       "R-201_Write_TO_T-101_DB".Abort := "R-201_SEQ_DB".S_NO >= 21 AND "R-201_SEQ_DB".S_NO <= 39;
       "R-201_Write_TO_T-102_DB".Abort := "R-201_SEQ_DB".S_NO >= 21 AND "R-201_SEQ_DB".S_NO <= 39;
       "R-201_Write_TO_T-103_DB".Abort :=("R-201_DB".Status.State = 3);

   END_IF;

   //***************Interlocks to T-104***************//
   "R-201_Write_TO_T-104_DB".ReqWater := "XV-2013_DB".CS AND "XV-1043_DB".OS AND ("R-201_DB".Status.Step = 23 OR "R-201_DB".Status.Step = 68 OR "R-201_DB".Status.Step = 66);

   //***************Valves Status***************//
   "R-201_Aux_DB"."Bool".TOff := "R-201_DB".Equipments.Valves."XV-2013".TurningOff OR "R-201_DB".Equipments.Valves."XV-2011".TurningOff OR "R-201_DB".Equipments.Valves."XV-2021".TurningOff OR "R-201_DB".Equipments.Valves."XV-1043".TurningOff;

   //***************Timers***************//
   //Pre-Mix Timer
   "R-201_Aux_DB"."Bool".PreMixT_En := "R-201_DB".Status.Step = 26 AND "R-201_Read_FROM_T-102_DB".Recirculating AND "R-201_Read_FROM_T-101_DB".Recirculating; //T-102 AND T-102 Mixing
   "R-201_Aux_DB"."Bool".PreMixT_Reset := "R-201_DB".Cmds.Abort OR "R-201_DB".Status.Step = 1;
   //pH Stabilize Timer
   "R-201_Aux_DB"."Bool".StabpHTEn := "R-201_Aux_DB"."Bool".StabpHTEnStep AND "FT-1021_DB".SAI > 0.1 AND "FT-1011_DB".SAI > 0.1;
   "R-201_Aux_DB"."Bool".StabpHTEn_Reset := "R-201_DB".Cmds.Abort OR "R-201_DB".Status.Step = 1;
   //Reaction Timer
   "R-201_Aux_DB"."Bool".ReactorTEn := "R-201_DB".Status.Step = 40;
   "R-201_Aux_DB"."Bool".ReactorT_Reset := "R-201_DB".Cmds.Abort OR "R-201_DB".Status.Step = 1;
   //Last Run Timer
   "R-201_Aux_DB"."Bool".FlushOutTEn := ("R-201_DB".Status.Step = 67 OR "R-201_DB".Status.Step = 64) AND ("P-201A_DB".CF OR "P-201B_DB".CF) AND "XV-2013_DB".OS;
   //Mix To Clean Timer
   "R-201_Aux_DB"."Bool".MixToCleanTEn := "R-201_DB".Status.Step = 63 AND "VFD-R201_DB".RUN_FEEDBACK;
   "R-201_Aux_DB"."Bool".MixToCleanT_Reset := "R-201_DB".Cmds.Abort OR "R-201_DB".Status.Step = 1;
END_FUNCTION

FUNCTION "R-201_SEQ_FC" : Void   // FC37, LAD
{ S7_Optimized_Access := 'TRUE' }
VERSION : 0.1
   VAR_TEMP   // added for the SCL form of the ladder/FBD networks
      _w1 : Bool;
      _w2 : Bool;
   END_VAR
BEGIN

REGION Network 2: Abort
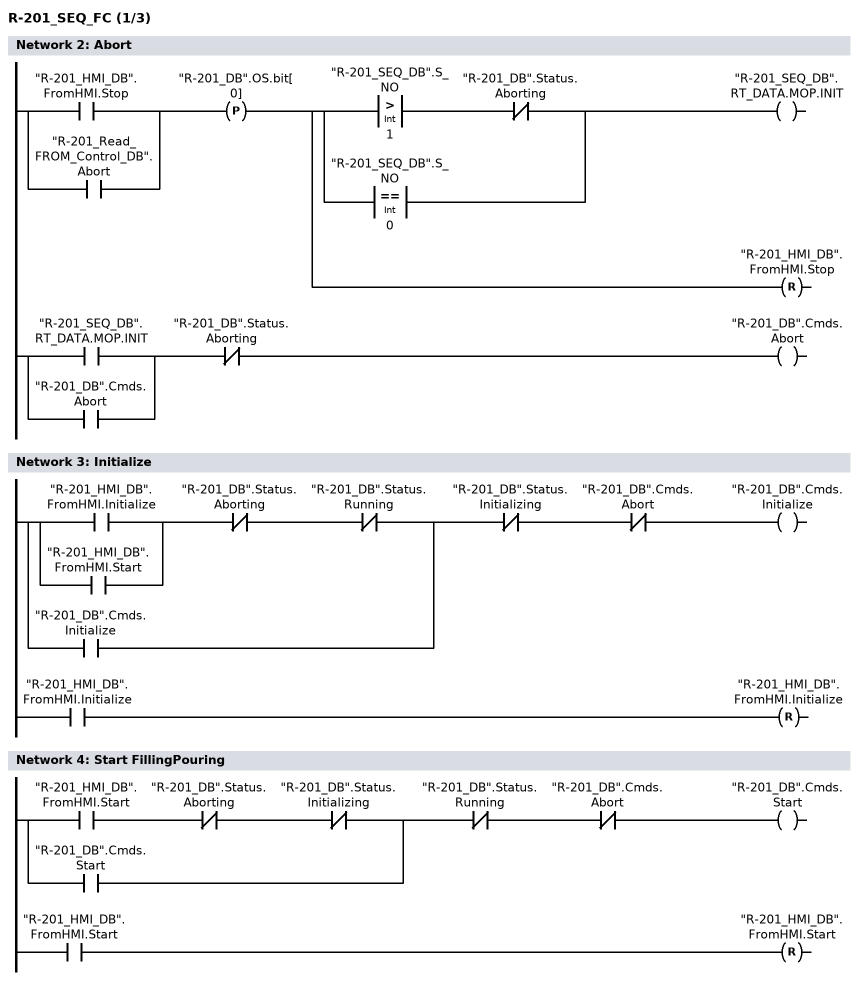
   RUNG wire#powerrail
      Contact( "R-201_HMI_DB".FromHMI.Stop )
      wire#w1
      P_Trig( "R-201_DB".OS.bit[0] )
      wire#w2
      { S7_Templates := "SrcType := Int" } GT_Contact(in1 := "R-201_SEQ_DB".S_NO, in2 := 1)
      I_Contact( "R-201_DB".Status.Aborting )
      wire#w3
      Coil( "R-201_SEQ_DB".RT_DATA.MOP.INIT )
   END_RUNG
   RUNG wire#powerrail
      Contact( "R-201_Read_FROM_Control_DB".Abort )
   END_RUNG wire#w1
   RUNG wire#w2
      { S7_Templates := "SrcType := Int" } EQ_Contact(in1 := "R-201_SEQ_DB".S_NO, in2 := 0)
   END_RUNG wire#w3
   RUNG wire#w2
      R_Coil( "R-201_HMI_DB".FromHMI.Stop )
   END_RUNG
   RUNG wire#powerrail
      Contact( "R-201_SEQ_DB".RT_DATA.MOP.INIT )
      wire#w4
      I_Contact( "R-201_DB".Status.Aborting )
      Coil( "R-201_DB".Cmds.Abort )
   END_RUNG
   RUNG wire#powerrail
      Contact( "R-201_DB".Cmds.Abort )
   END_RUNG wire#w4
   // the same network as SCL:
   #_w1 := "R-201_HMI_DB".FromHMI.Stop OR "R-201_Read_FROM_Control_DB".Abort;
   #_w2 := #_w1 AND NOT "R-201_DB".OS.bit[0];   // rising edge
   "R-201_DB".OS.bit[0] := #_w1;
   "R-201_SEQ_DB".RT_DATA.MOP.INIT := #_w2 AND ((("R-201_SEQ_DB".S_NO > 1) AND NOT "R-201_DB".Status.Aborting) OR ("R-201_SEQ_DB".S_NO = 0));
   IF #_w2 THEN "R-201_HMI_DB".FromHMI.Stop := FALSE; END_IF;
   "R-201_DB".Cmds.Abort := ("R-201_SEQ_DB".RT_DATA.MOP.INIT OR "R-201_DB".Cmds.Abort) AND NOT "R-201_DB".Status.Aborting;
END_REGION

REGION Network 3: Initialize
   RUNG wire#powerrail
      Contact( "R-201_HMI_DB".FromHMI.Initialize )
      wire#w1
      I_Contact( "R-201_DB".Status.Aborting )
      I_Contact( "R-201_DB".Status.Running )
      wire#w2
      I_Contact( "R-201_DB".Status.Initializing )
      I_Contact( "R-201_DB".Cmds.Abort )
      Coil( "R-201_DB".Cmds.Initialize )
   END_RUNG
   RUNG wire#powerrail
      Contact( "R-201_HMI_DB".FromHMI.Start )
   END_RUNG wire#w1
   RUNG wire#powerrail
      Contact( "R-201_DB".Cmds.Initialize )
   END_RUNG wire#w2
   RUNG wire#powerrail
      Contact( "R-201_HMI_DB".FromHMI.Initialize )
      R_Coil( "R-201_HMI_DB".FromHMI.Initialize )
   END_RUNG
   // the same network as SCL:
   "R-201_DB".Cmds.Initialize := ((("R-201_HMI_DB".FromHMI.Initialize OR "R-201_HMI_DB".FromHMI.Start) AND NOT "R-201_DB".Status.Aborting AND NOT "R-201_DB".Status.Running) OR "R-201_DB".Cmds.Initialize) AND NOT "R-201_DB".Status.Initializing AND NOT "R-201_DB".Cmds.Abort;
   IF "R-201_HMI_DB".FromHMI.Initialize THEN "R-201_HMI_DB".FromHMI.Initialize := FALSE; END_IF;
END_REGION

REGION Network 4: Start FillingPouring
   RUNG wire#powerrail
      Contact( "R-201_HMI_DB".FromHMI.Start )
      I_Contact( "R-201_DB".Status.Aborting )
      I_Contact( "R-201_DB".Status.Initializing )
      wire#w1
      I_Contact( "R-201_DB".Status.Running )
      I_Contact( "R-201_DB".Cmds.Abort )
      Coil( "R-201_DB".Cmds.Start )
   END_RUNG
   RUNG wire#powerrail
      Contact( "R-201_DB".Cmds.Start )
   END_RUNG wire#w1
   RUNG wire#powerrail
      Contact( "R-201_HMI_DB".FromHMI.Start )
      R_Coil( "R-201_HMI_DB".FromHMI.Start )
   END_RUNG
   // the same network as SCL:
   "R-201_DB".Cmds.Start := (("R-201_HMI_DB".FromHMI.Start AND NOT "R-201_DB".Status.Aborting AND NOT "R-201_DB".Status.Initializing) OR "R-201_DB".Cmds.Start) AND NOT "R-201_DB".Status.Running AND NOT "R-201_DB".Cmds.Abort;
   IF "R-201_HMI_DB".FromHMI.Start THEN "R-201_HMI_DB".FromHMI.Start := FALSE; END_IF;
END_REGION

REGION Network 5: Procedure Selected
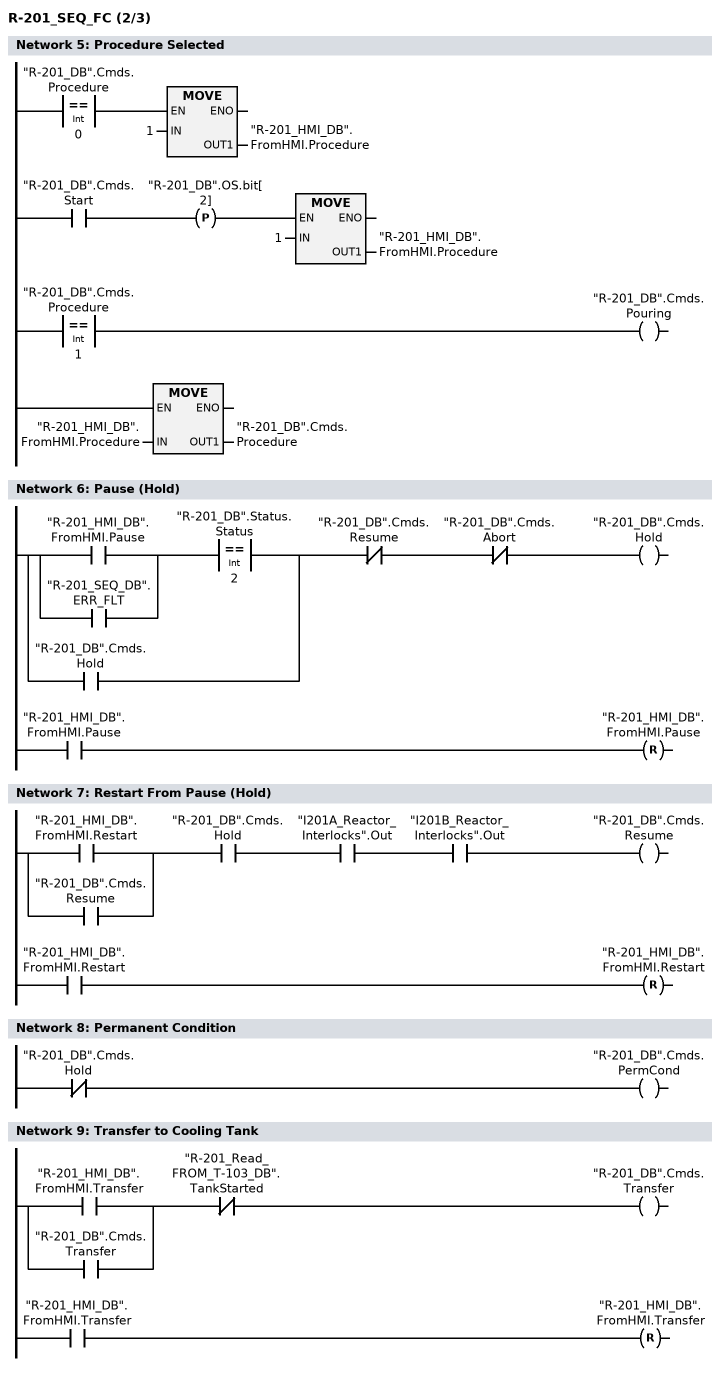
   RUNG wire#powerrail
      { S7_Templates := "SrcType := Int" } EQ_Contact(in1 := "R-201_DB".Cmds.Procedure, in2 := 0)
      Move(in := 1, out1 => "R-201_HMI_DB".FromHMI.Procedure)
   END_RUNG
   RUNG wire#powerrail
      Contact( "R-201_DB".Cmds.Start )
      P_Trig( "R-201_DB".OS.bit[2] )
      Move(in := 1, out1 => "R-201_HMI_DB".FromHMI.Procedure)
   END_RUNG
   RUNG wire#powerrail
      { S7_Templates := "SrcType := Int" } EQ_Contact(in1 := "R-201_DB".Cmds.Procedure, in2 := 1)
      Coil( "R-201_DB".Cmds.Pouring )
   END_RUNG
   RUNG wire#powerrail
      Move(in := "R-201_HMI_DB".FromHMI.Procedure, out1 => "R-201_DB".Cmds.Procedure)
   END_RUNG
   // the same network as SCL:
   IF "R-201_DB".Cmds.Procedure = 0 THEN "R-201_HMI_DB".FromHMI.Procedure := 1; END_IF;
   #_w1 := "R-201_DB".Cmds.Start AND NOT "R-201_DB".OS.bit[2];   // rising edge
   "R-201_DB".OS.bit[2] := "R-201_DB".Cmds.Start;
   IF #_w1 THEN "R-201_HMI_DB".FromHMI.Procedure := 1; END_IF;
   "R-201_DB".Cmds.Pouring := "R-201_DB".Cmds.Procedure = 1;
   "R-201_DB".Cmds.Procedure := "R-201_HMI_DB".FromHMI.Procedure;
END_REGION

REGION Network 6: Pause (Hold)
   RUNG wire#powerrail
      Contact( "R-201_HMI_DB".FromHMI.Pause )
      wire#w1
      { S7_Templates := "SrcType := Int" } EQ_Contact(in1 := "R-201_DB".Status.Status, in2 := 2)
      wire#w2
      I_Contact( "R-201_DB".Cmds.Resume )
      I_Contact( "R-201_DB".Cmds.Abort )
      Coil( "R-201_DB".Cmds.Hold )
   END_RUNG
   RUNG wire#powerrail
      Contact( "R-201_SEQ_DB".ERR_FLT )
   END_RUNG wire#w1
   RUNG wire#powerrail
      Contact( "R-201_DB".Cmds.Hold )
   END_RUNG wire#w2
   RUNG wire#powerrail
      Contact( "R-201_HMI_DB".FromHMI.Pause )
      R_Coil( "R-201_HMI_DB".FromHMI.Pause )
   END_RUNG
   // the same network as SCL:
   "R-201_DB".Cmds.Hold := ((("R-201_HMI_DB".FromHMI.Pause OR "R-201_SEQ_DB".ERR_FLT) AND ("R-201_DB".Status.Status = 2)) OR "R-201_DB".Cmds.Hold) AND NOT "R-201_DB".Cmds.Resume AND NOT "R-201_DB".Cmds.Abort;
   IF "R-201_HMI_DB".FromHMI.Pause THEN "R-201_HMI_DB".FromHMI.Pause := FALSE; END_IF;
END_REGION

REGION Network 7: Restart From Pause (Hold)
   RUNG wire#powerrail
      Contact( "R-201_HMI_DB".FromHMI.Restart )
      wire#w1
      Contact( "R-201_DB".Cmds.Hold )
      Contact( "I201A_Reactor_Interlocks".Out )
      Contact( "I201B_Reactor_Interlocks".Out )
      Coil( "R-201_DB".Cmds.Resume )
   END_RUNG
   RUNG wire#powerrail
      Contact( "R-201_DB".Cmds.Resume )
   END_RUNG wire#w1
   RUNG wire#powerrail
      Contact( "R-201_HMI_DB".FromHMI.Restart )
      R_Coil( "R-201_HMI_DB".FromHMI.Restart )
   END_RUNG
   // the same network as SCL:
   "R-201_DB".Cmds.Resume := ("R-201_HMI_DB".FromHMI.Restart OR "R-201_DB".Cmds.Resume) AND "R-201_DB".Cmds.Hold AND "I201A_Reactor_Interlocks".Out AND "I201B_Reactor_Interlocks".Out;
   IF "R-201_HMI_DB".FromHMI.Restart THEN "R-201_HMI_DB".FromHMI.Restart := FALSE; END_IF;
END_REGION

REGION Network 8: Permanent Condition
   RUNG wire#powerrail
      I_Contact( "R-201_DB".Cmds.Hold )
      Coil( "R-201_DB".Cmds.PermCond )
   END_RUNG
   // the same network as SCL:
   "R-201_DB".Cmds.PermCond := NOT "R-201_DB".Cmds.Hold;
END_REGION

REGION Network 9: Transfer to Cooling Tank
   RUNG wire#powerrail
      Contact( "R-201_HMI_DB".FromHMI.Transfer )
      wire#w1
      I_Contact( "R-201_Read_FROM_T-103_DB".TankStarted )
      Coil( "R-201_DB".Cmds.Transfer )
   END_RUNG
   RUNG wire#powerrail
      Contact( "R-201_DB".Cmds.Transfer )
   END_RUNG wire#w1
   RUNG wire#powerrail
      Contact( "R-201_HMI_DB".FromHMI.Transfer )
      R_Coil( "R-201_HMI_DB".FromHMI.Transfer )
   END_RUNG
   // the same network as SCL:
   "R-201_DB".Cmds.Transfer := ("R-201_HMI_DB".FromHMI.Transfer OR "R-201_DB".Cmds.Transfer) AND NOT "R-201_Read_FROM_T-103_DB".TankStarted;
   IF "R-201_HMI_DB".FromHMI.Transfer THEN "R-201_HMI_DB".FromHMI.Transfer := FALSE; END_IF;
END_REGION

REGION Network 10: Tank Wash
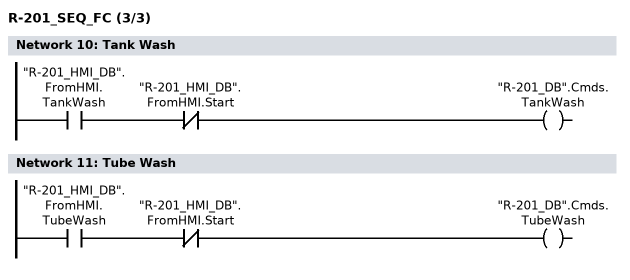
   RUNG wire#powerrail
      Contact( "R-201_HMI_DB".FromHMI.TankWash )
      I_Contact( "R-201_HMI_DB".FromHMI.Start )
      Coil( "R-201_DB".Cmds.TankWash )
   END_RUNG
   // the same network as SCL:
   "R-201_DB".Cmds.TankWash := "R-201_HMI_DB".FromHMI.TankWash AND NOT "R-201_HMI_DB".FromHMI.Start;
END_REGION

REGION Network 11: Tube Wash
   RUNG wire#powerrail
      Contact( "R-201_HMI_DB".FromHMI.TubeWash )
      I_Contact( "R-201_HMI_DB".FromHMI.Start )
      Coil( "R-201_DB".Cmds.TubeWash )
   END_RUNG
   // the same network as SCL:
   "R-201_DB".Cmds.TubeWash := "R-201_HMI_DB".FromHMI.TubeWash AND NOT "R-201_HMI_DB".FromHMI.Start;
END_REGION

REGION Network 12 (SCL): Sequence Status
   IF "R-201_SEQ_DB".S_NO = 1 THEN
       "R-201_DB".Status.Status := 1; //Idle
   ELSIF ("R-201_SEQ_DB".S_NO > 1 AND "R-201_SEQ_DB".S_NO <= 150)  AND NOT "R-201_SEQ_DB".ERR_FLT AND NOT "R-201_DB".Cmds.Hold THEN
       "R-201_DB".Status.Status := 2; //Running
   ELSIF "R-201_SEQ_DB".S_NO >= 151 AND "R-201_SEQ_DB".S_NO <= 160 AND NOT "R-201_SEQ_DB".ERR_FLT THEN
       "R-201_DB".Status.Status := 3; // Stopping
   ELSIF "R-201_SEQ_DB".ERR_FLT  AND ("R-201_SEQ_DB".S_NO > 1 AND "R-201_SEQ_DB".S_NO <= 150) THEN
       "R-201_DB".Status.Status := 4; //Held
   ELSIF "R-201_SEQ_DB".ERR_FLT AND  ("R-201_SEQ_DB".S_NO > 1 AND "R-201_SEQ_DB".S_NO <= 150) AND "R-201_Aux_DB"."Bool".TOff  THEN
       "R-201_DB".Status.Status := 5; // Holding
   ELSE
       "R-201_DB".Status.Status := 6; // Unknown
   END_IF;


   "R-201_DB".Status.Running := ("R-201_SEQ_DB".S_NO > 3 AND "R-201_SEQ_DB".S_NO <= 150);
   "R-201_DB".Status.Initializing := ("R-201_SEQ_DB".S_NO >= 141 AND "R-201_SEQ_DB".S_NO <= 150);
   //Enable/Disable HMI Start/Stop Button
   "R-201_HMI_DB".ToHMI.EnStopButton:=("R-201_DB".Status.Status>1) OR "R-201_DB".Status.Step=0; //Enable HMI Stop Button
   "R-201_HMI_DB".ToHMI.EnStartButton:= "R-201_DB".Status.Status = 1; //Enable Start Button
   "R-201_HMI_DB".ToHMI.EnPauseButton := "R-201_DB".Status.Status = 2; //Enable Pause Button
   "R-201_HMI_DB".ToHMI.EnRestartButton := "R-201_DB".Status.Status = 4; //Enable Restart Button

   //****Interlock Activated
   "R-201_HMI_DB".ToHMI.InterlockActivated := "I201A_Reactor_Interlocks".Out AND "I201B_Reactor_Interlocks".Out;
END_REGION

REGION Network 13 (SCL): Sequence Step
   "R-201_DB".Status.Step := "R-201_SEQ_DB".S_NO;
END_REGION

REGION Network 14 (SCL): Sequence state (Procedure running)
   IF "R-201_SEQ_DB".S_NO = 3 OR "R-201_SEQ_DB".S_NO = 4 THEN
       "R-201_DB".Status.State := 1; //Seq Selection
   ELSIF "R-201_SEQ_DB".S_NO >= 21 AND "R-201_SEQ_DB".S_NO <= 60 THEN
       "R-201_DB".Status.State := 2; //Pouring 
   ELSIF "R-201_SEQ_DB".S_NO >= 61 AND "R-201_SEQ_DB".S_NO <= 80 THEN
       "R-201_DB".Status.State := 3; //Transfering
   ELSIF "R-201_SEQ_DB".S_NO >= 81 AND "R-201_SEQ_DB".S_NO <= 100 THEN
       "R-201_DB".Status.State := 4; //Washing Tank
   ELSIF "R-201_SEQ_DB".S_NO >= 101 AND "R-201_SEQ_DB".S_NO <= 140 THEN
       "R-201_DB".Status.State := 5; //Washing Lines
   ELSIF "R-201_SEQ_DB".S_NO >= 151 AND "R-201_SEQ_DB".S_NO <= 160 THEN
       "R-201_DB".Status.State := 6; //Aborting
   ELSIF "R-201_SEQ_DB".S_NO >= 141 AND "R-201_SEQ_DB".S_NO <= 150 THEN
       "R-201_DB".Status.State := 7; //Initializing
   ELSE
       "R-201_DB".Status.State := 0;
   END_IF;
END_REGION
END_FUNCTION

FUNCTION "R-201_Transitions_FC" : Void   // FC42, SCL
{ S7_Optimized_Access := 'TRUE' }
VERSION : 0.1
BEGIN

   //*****"Transition" for Low Level and Low pressure meaning "Tank is Empty"
   "R-201_Aux_DB"."Bool".Transitions.TankEmpty := "LT-2011_DB".SAI <= "ReactorLowLevelSetpoint" AND (("PT-201A_DB".SAI <= 1.0) AND ("PT-201B_DB".SAI <= 1.0));
END_FUNCTION

// folder: State MACHINE/2)Reactors/Reactor R-201/Control R-201

FUNCTION_BLOCK "R-201_Control"   // FB36, GRAPH_PLUS
{ S7_Optimized_Access := 'TRUE' }
VERSION : 0.1
   VAR_INPUT
      OFF_SQ : Bool := false;   // Turn sequence off
      INIT_SQ : Bool := false;   // Set sequence to initial state
      ACK_EF : Bool := false;   // Acknowledge all errors and faults
      "P-201A/B _SEL" : Int := 1;   // IF FALSE P201A is priority / IF TRUE P201B is priority
      "P-202A/B _SEL" : Int := 1;   // IF FALSE P202A is priority / IF TRUE P202B is priority
      IL : Bool;   // INTERLOCKS
   END_VAR
   VAR_OUTPUT
      S_NO : Int := 0;   // Step number
      S_MORE : Bool := false;   // More steps are available and can be shown in S_NO
      S_ACTIVE : Bool := false;   // Step indicated in S_NO is active
      ERR_FLT : Bool := false;   // Interlock or supervision group error
      AUTO_ON : Bool := false;   // Automatic mode is active
   END_VAR
   VAR
      STATE : Int;   // Step number
      Reactor : Struct
         ABORTING : Bool;   // Sequence about
         BatchVolume : Real;   // Batch Volume SP in Liter
         Batchsize : Real;   // Batch size in SP Liter
      END_STRUCT;
      TEMP : Struct
         TANKS_BATCH : Real;   // T-101 & T-102 Batch Sizes
         "EMPTY_LV_0%" : Real;   // 0 % of the Total Batch Size SP
         "MIN_LV_20%" : Real;   // 20 % of the Total Batch Size SP
         "MAX_LV_80%" : Real;   // 80 % of the Total Batch Size SP
         "BELOW_32%" : Real;   // <32% of T-103 Total Batch Size
         "Greater_8%" : Real;   // >8% of T-103 Total Batch Size
         "PRE-ADD" : Real;   // Water & Batch size
         X_SOL_SIZE : Real := 5.0;   // T-101 Soluction Size
         Y_SOL_SIZE : Real := 5.0;   // T-102 Soluction Size
         OFFSEt : Struct
            MAX : Real;
            MIN : Real;
         END_STRUCT;
      END_STRUCT;
      "R-202_TEMP" : Struct
         TANKS_BATCH : Real;   // T-101 & T-102 Batch Sizes
         "EMPTY_LV_0%" : Real;   // 0 % of the Total Batch Size SP
         "MIN_LV_20%" : Real;   // 20 % of the Total Batch Size SP
         "MAX_LV_80%" : Real;   // 80 % of the Total Batch Size SP
         "BELOW_32%" : Real;   // <32% of T-103 Total Batch Size
         "Greater_8%" : Real;   // >8% of T-103 Total Batch Size
         "PRE-ADD" : Real;   // Water & Batch size
         X_SOL_SIZE : Real := 5.0;   // T-101 Soluction Size
         Y_SOL_SIZE : Real := 5.0;   // T-102 Soluction Size
         OFFSEt : Struct
            MAX : Real;
            MIN : Real;
         END_STRUCT;
      END_STRUCT;
      "TIMER" : Array[0..10] of IEC_TIMER;
      "TIME" : Array[0..10] of Time;
      HMI_INFO : Array[0..12] of UInt;
      IF_PAR : G7_IfParPlus_V6;
      RT_DATA : G7_RTDataPlus_V6;   // Internal data area
      Abort : G7_TransitionPlus_V6;   // Transition structure
      "Init R-201" : G7_TransitionPlus_V6;   // Transition structure
      RProcess : G7_TransitionPlus_V6;   // Transition structure
      Trans14 : G7_TransitionPlus_V6;   // Transition structure
      Trans105 : G7_TransitionPlus_V6;   // Transition structure
      Trans106 : G7_TransitionPlus_V6;   // Transition structure
      BachSize : G7_TransitionPlus_V6;   // Transition structure
      Trans110 : G7_TransitionPlus_V6;   // Transition structure
      Trans111 : G7_TransitionPlus_V6;   // Transition structure
      PresetsOK : G7_TransitionPlus_V6;   // Transition structure
      FromHMI : G7_TransitionPlus_V6;   // Transition structure
      Started : G7_TransitionPlus_V6;   // Transition structure
      RDone : G7_TransitionPlus_V6;   // Transition structure
      TDone : G7_TransitionPlus_V6;   // Transition structure
      "R-201 Idle" : G7_TransitionPlus_V6;   // Transition structure
      Trans19 : G7_TransitionPlus_V6;   // Transition structure
      TaW : G7_TransitionPlus_V6;   // Transition structure
      TuW : G7_TransitionPlus_V6;   // Transition structure
      Trans21 : G7_TransitionPlus_V6;   // Transition structure
      DoneAbrt : G7_TransitionPlus_V6;   // Transition structure
      "R-201_Idle" : G7_TransitionPlus_V6;   // Transition structure
      Trans116 : G7_TransitionPlus_V6;   // Transition structure
      Trans117 : G7_TransitionPlus_V6;   // Transition structure
      Trans118 : G7_TransitionPlus_V6;   // Transition structure
      Trans119 : G7_TransitionPlus_V6;   // Transition structure
      Idle : G7_StepPlus_V6;   // Step structure
      Initialize : G7_StepPlus_V6;   // Step structure
      Ready : G7_StepPlus_V6;   // Step structure
      TankWash : G7_StepPlus_V6;   // Step structure
      TubingWash : G7_StepPlus_V6;   // Step structure
      Bach_Size : G7_StepPlus_V6;   // Step structure
      Presets : G7_StepPlus_V6;   // Step structure
      WaitHMI : G7_StepPlus_V6;   // Step structure
      Start : G7_StepPlus_V6;   // Step structure
      Reacting : G7_StepPlus_V6;   // Step structure
      "Transf-->T-103" : G7_StepPlus_V6;   // Step structure
      DoneTransfer : G7_StepPlus_V6;   // Step structure
      Aborting : G7_StepPlus_V6;   // Step structure
      Release : G7_StepPlus_V6;   // Step structure
      WaterIn : G7_StepPlus_V6;   // Step structure
      Release_TW : G7_StepPlus_V6;   // Step structure
      Release_TuW : G7_StepPlus_V6;   // Step structure
      RdyTaW : G7_StepPlus_V6;   // Step structure
      Wait : G7_StepPlus_V6;   // Step structure
      RdyTuW : G7_StepPlus_V6;   // Step structure
      Pouring_X_Y : G7_StepPlus_V6;   // Step structure
      WaitTransfer : G7_StepPlus_V6;   // Step structure
      SINI : Array[0..5] of USInt;
      LSTT : Array[0..24] of USInt;
      ATAJ : Array[0..24] of USInt;
      ATAB : Array[0..24] of USInt;
      PSTT : Array[0..24] of USInt;
      NSTT : Array[0..24] of USInt;
      ASSJ : Array[0..21] of USInt;
      ASSB : Array[0..21] of USInt;
      PTTS : Array[0..21] of USInt;
      NTTS : Array[0..21] of USInt;
      SW_SQTS : Array[0..21] of USInt;
      SWITCH : Array[0..4] of USInt;
      TVX : Array[0..10] of USInt;
      TTX : Array[0..10] of USInt;
      TSX : Array[0..5] of USInt;
      S00X : Array[0..5] of USInt;
      SOFFX : Array[0..5] of USInt;
      SONX : Array[0..5] of USInt;
      SAX : Array[0..5] of USInt;
      SERRX : Array[0..22] of USInt;
      SMX : Array[0..22] of USInt;
      S0X : Array[0..22] of USInt;
      S1X : Array[0..22] of USInt;
      IL_ALARM_INST : Diag_Alarm;
      SUP_ALARM_INST : Diag_Alarm;
      STEP_TIME_ALARM_INST : Diag_Alarm;
      IEC_TIMER_INST : IEC_TIMER;
      TRANSACTION_FLAG : Bool := false;
   END_VAR
   VAR CONSTANT
      "Single R-201 T-101 seq done" : Int := 214;
      "Single R-201 T-102 seq done" : Int := 218;
   END_VAR
   // SINI[0] := 2;
   // LSTT[0] := 12;
   // NSTT[0] := 12;
   // PTTS[0] := 255;
   // TVX[0] := 16#1;
   // TTX[0] := 16#1;
   // TSX[0] := 16#1;
   // S00X[0] := 16#1;
   // SOFFX[0] := 16#1;
   // SONX[0] := 16#1;
   // SAX[0] := 16#1;
   // SERRX[0] := 16#1;
   // SMX[0] := 16#1;
   // S0X[0] := 16#1;
   // S1X[0] := 16#1;
   // SINI[2] := 255;
   // SINI[3] := 255;
   // SINI[4] := 255;
   // SINI[5] := 255;
   // LSTT[1] := 255;
   // LSTT[2] := 2;
   // LSTT[3] := 255;
   // LSTT[4] := 255;
   // LSTT[5] := 255;
   // LSTT[6] := 255;
   // LSTT[19] := 255;
   // LSTT[9] := 255;
   // LSTT[10] := 255;
   // LSTT[11] := 255;
   // LSTT[12] := 255;
   // LSTT[13] := 255;
   // LSTT[18] := 255;
   // LSTT[15] := 255;
   // LSTT[16] := 17;
   // LSTT[17] := 19;
   // LSTT[21] := 255;
   // LSTT[22] := 255;
   // LSTT[23] := 255;
   // LSTT[24] := 255;
   // ATAJ[1] := 1;
   // ATAJ[2] := 2;
   // ATAJ[3] := 3;
   // ATAJ[4] := 4;
   // ATAJ[5] := 5;
   // ATAJ[6] := 6;
   // ATAJ[7] := 7;
   // ATAJ[8] := 8;
   // ATAJ[9] := 9;
   // ATAJ[10] := 10;
   // ATAJ[11] := 11;
   // ATAJ[12] := 12;
   // ATAJ[13] := 13;
   // ATAJ[14] := 14;
   // ATAJ[15] := 15;
   // ATAJ[16] := 16;
   // ATAJ[17] := 17;
   // ATAJ[18] := 18;
   // ATAJ[19] := 19;
   // ATAJ[20] := 20;
   // ATAJ[21] := 21;
   // ATAJ[22] := 22;
   // ATAJ[23] := 23;
   // ATAJ[24] := 24;
   // ATAB[20] := 20;
   // ATAB[2] := 16;
   // ATAB[3] := 3;
   // ATAB[4] := 4;
   // ATAB[5] := 5;
   // ATAB[6] := 6;
   // ATAB[7] := 7;
   // ATAB[8] := 8;
   // ATAB[9] := 9;
   // ATAB[10] := 10;
   // ATAB[11] := 11;
   // ATAB[12] := 12;
   // ATAB[13] := 13;
   // ATAB[14] := 14;
   // ATAB[15] := 15;
   // ATAB[16] := 17;
   // ATAB[17] := 2;
   // ATAB[18] := 18;
   // ATAB[19] := 19;
   // ATAB[21] := 21;
   // ATAB[22] := 22;
   // ATAB[23] := 23;
   // ATAB[24] := 24;
   // PSTT[20] := 13;
   // PSTT[2] := 1;
   // PSTT[3] := 2;
   // PSTT[4] := 3;
   // PSTT[5] := 4;
   // PSTT[6] := 5;
   // PSTT[7] := 15;
   // PSTT[8] := 16;
   // PSTT[9] := 6;
   // PSTT[10] := 7;
   // PSTT[11] := 8;
   // PSTT[12] := 9;
   // PSTT[13] := 10;
   // PSTT[14] := 11;
   // PSTT[15] := 17;
   // PSTT[16] := 1;
   // PSTT[17] := 1;
   // PSTT[18] := 19;
   // PSTT[19] := 12;
   // PSTT[21] := 14;
   // PSTT[22] := 20;
   // PSTT[23] := 18;
   // PSTT[24] := 21;
   // NSTT[1] := 1;
   // NSTT[2] := 2;
   // NSTT[3] := 5;
   // NSTT[4] := 15;
   // NSTT[5] := 16;
   // NSTT[6] := 6;
   // NSTT[19] := 13;
   // NSTT[9] := 7;
   // NSTT[10] := 8;
   // NSTT[11] := 14;
   // NSTT[12] := 21;
   // NSTT[13] := 11;
   // NSTT[18] := 4;
   // NSTT[15] := 3;
   // NSTT[16] := 17;
   // NSTT[17] := 19;
   // NSTT[21] := 18;
   // NSTT[22] := 9;
   // NSTT[23] := 20;
   // NSTT[24] := 10;
   // ASSJ[1] := 1;
   // ASSJ[2] := 2;
   // ASSJ[3] := 3;
   // ASSJ[4] := 4;
   // ASSJ[5] := 5;
   // ASSJ[6] := 6;
   // ASSJ[7] := 7;
   // ASSJ[8] := 8;
   // ASSJ[9] := 9;
   // ASSJ[10] := 10;
   // ASSJ[11] := 11;
   // ASSJ[12] := 12;
   // ASSJ[13] := 13;
   // ASSJ[14] := 14;
   // ASSJ[15] := 15;
   // ASSJ[16] := 16;
   // ASSJ[17] := 17;
   // ASSJ[18] := 18;
   // ASSJ[19] := 19;
   // ASSJ[20] := 20;
   // ASSJ[21] := 21;
   // ASSB[1] := 1;
   // ASSB[2] := 2;
   // ASSB[3] := 3;
   // ASSB[4] := 4;
   // ASSB[5] := 5;
   // ASSB[6] := 6;
   // ASSB[7] := 7;
   // ASSB[8] := 8;
   // ASSB[9] := 9;
   // ASSB[10] := 10;
   // ASSB[11] := 11;
   // ASSB[12] := 12;
   // ASSB[13] := 13;
   // ASSB[14] := 14;
   // ASSB[15] := 15;
   // ASSB[16] := 16;
   // ASSB[17] := 17;
   // ASSB[18] := 18;
   // ASSB[19] := 19;
   // ASSB[20] := 20;
   // ASSB[21] := 21;
   // PTTS[2] := 255;
   // PTTS[3] := 15;
   // PTTS[4] := 18;
   // PTTS[5] := 3;
   // PTTS[6] := 6;
   // PTTS[7] := 9;
   // PTTS[8] := 10;
   // PTTS[9] := 22;
   // PTTS[10] := 24;
   // PTTS[11] := 13;
   // PTTS[12] := 255;
   // PTTS[13] := 19;
   // PTTS[14] := 11;
   // PTTS[16] := 5;
   // PTTS[17] := 255;
   // PTTS[18] := 21;
   // PTTS[19] := 255;
   // PTTS[20] := 23;
   // PTTS[21] := 12;
   // PTTS[15] := 4;
   // NTTS[1] := 2;
   // NTTS[2] := 3;
   // NTTS[3] := 4;
   // NTTS[4] := 5;
   // NTTS[5] := 6;
   // NTTS[6] := 9;
   // NTTS[7] := 10;
   // NTTS[8] := 11;
   // NTTS[9] := 12;
   // NTTS[10] := 13;
   // NTTS[11] := 14;
   // NTTS[12] := 19;
   // NTTS[13] := 20;
   // NTTS[14] := 21;
   // NTTS[15] := 7;
   // NTTS[16] := 8;
   // NTTS[17] := 15;
   // NTTS[18] := 23;
   // NTTS[19] := 18;
   // NTTS[20] := 22;
   // NTTS[21] := 24;
   // SW_SQTS[2] := 2;
   // SW_SQTS[3] := 3;
   // SW_SQTS[4] := 4;
   // SW_SQTS[5] := 2;
   // SW_SQTS[6] := 2;
   // SW_SQTS[7] := 2;
   // SW_SQTS[8] := 2;
   // SW_SQTS[9] := 2;
   // SW_SQTS[10] := 2;
   // SW_SQTS[11] := 2;
   // SW_SQTS[12] := 5;
   // SW_SQTS[13] := 5;
   // SW_SQTS[14] := 2;
   // SW_SQTS[15] := 3;
   // SW_SQTS[16] := 4;
   // SW_SQTS[17] := 3;
   // SW_SQTS[18] := 2;
   // SW_SQTS[19] := 4;
   // SW_SQTS[20] := 2;
   // SW_SQTS[21] := 2;
   // SWITCH[1] := 191;
   // SWITCH[2] := 223;
   // SWITCH[3] := 239;
   // SWITCH[4] := 7;
   // ATAB[0] := 1;
   // PTTS[1] := 1;
   // SW_SQTS[1] := 1;
   // SWITCH[0] := 60;
BEGIN
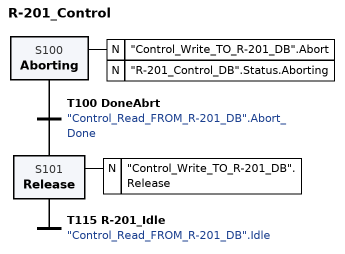
   // sequencer 1
   STEP Aborting:   // S100, max time T#10S, warning time T#7S
      // T-101 Pouring Soluction Valve
              N    "Control_Write_TO_R-201_DB".Abort
              N    "R-201_Control_DB".Status.Aborting
   END_STEP
   TRANSITION DoneAbrt FROM Aborting TO Release   // T100: CLOSED: XV-1041 XV-1011 XV-1013OFF: VFD-1011 P-101A P-101BZERO: FT-1041 Totalizer
      := "Control_Read_FROM_R-201_DB".Abort_Done;
   END_TRANSITION
   STEP Release:   // S101, max time T#10S, warning time T#7S
              N    "Control_Write_TO_R-201_DB".Release
   END_STEP
   TRANSITION "R-201_Idle" FROM Release TO ?   // T115
      := "Control_Read_FROM_R-201_DB".Idle;
   END_TRANSITION
END_FUNCTION_BLOCK

FUNCTION "R-201_CTRL_SEQ_FC" : Void   // FC38, LAD
{ S7_Optimized_Access := 'TRUE' }
VERSION : 0.1
   VAR_TEMP   // added for the SCL form of the ladder/FBD networks
      _w1 : Bool;
   END_VAR
BEGIN

REGION Network 2: Reset Abort Cmd
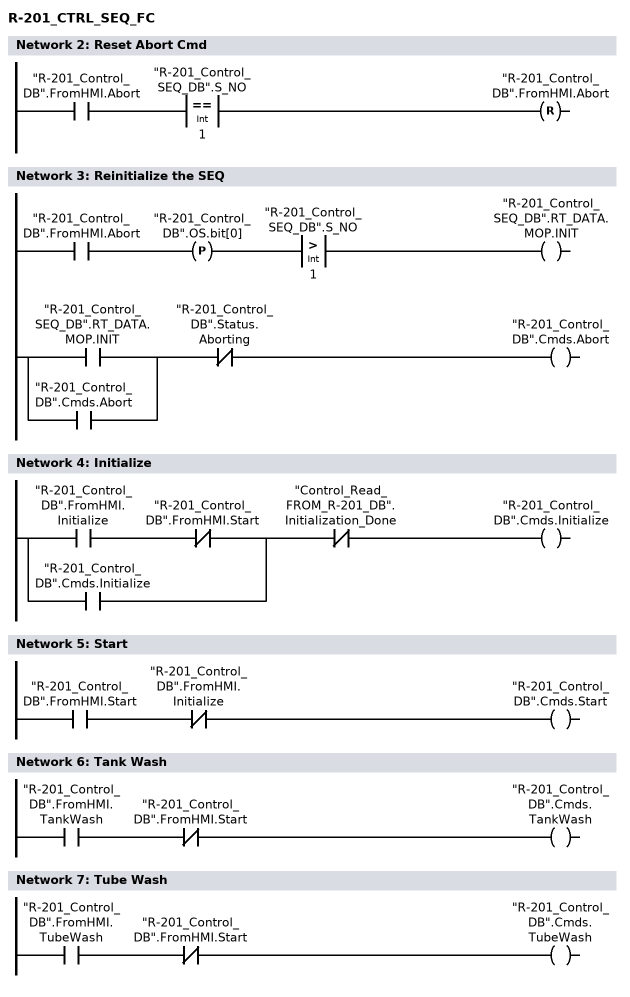
   RUNG wire#powerrail
      Contact( "R-201_Control_DB".FromHMI.Abort )
      { S7_Templates := "SrcType := Int" } EQ_Contact(in1 := "R-201_Control_SEQ_DB".S_NO, in2 := 1)
      R_Coil( "R-201_Control_DB".FromHMI.Abort )
   END_RUNG
   // the same network as SCL:
   IF "R-201_Control_DB".FromHMI.Abort AND ("R-201_Control_SEQ_DB".S_NO = 1) THEN
       "R-201_Control_DB".FromHMI.Abort := FALSE;
   END_IF;
END_REGION

REGION Network 3: Reinitialize the SEQ
   RUNG wire#powerrail
      Contact( "R-201_Control_DB".FromHMI.Abort )
      P_Trig( "R-201_Control_DB".OS.bit[0] )
      { S7_Templates := "SrcType := Int" } GT_Contact(in1 := "R-201_Control_SEQ_DB".S_NO, in2 := 1)
      Coil( "R-201_Control_SEQ_DB".RT_DATA.MOP.INIT )
   END_RUNG
   RUNG wire#powerrail
      Contact( "R-201_Control_SEQ_DB".RT_DATA.MOP.INIT )
      wire#w1
      I_Contact( "R-201_Control_DB".Status.Aborting )
      Coil( "R-201_Control_DB".Cmds.Abort )
   END_RUNG
   RUNG wire#powerrail
      Contact( "R-201_Control_DB".Cmds.Abort )
   END_RUNG wire#w1
   // the same network as SCL:
   #_w1 := "R-201_Control_DB".FromHMI.Abort AND NOT "R-201_Control_DB".OS.bit[0];   // rising edge
   "R-201_Control_DB".OS.bit[0] := "R-201_Control_DB".FromHMI.Abort;
   "R-201_Control_SEQ_DB".RT_DATA.MOP.INIT := #_w1 AND ("R-201_Control_SEQ_DB".S_NO > 1);
   "R-201_Control_DB".Cmds.Abort := ("R-201_Control_SEQ_DB".RT_DATA.MOP.INIT OR "R-201_Control_DB".Cmds.Abort) AND NOT "R-201_Control_DB".Status.Aborting;
END_REGION

REGION Network 4: Initialize
   RUNG wire#powerrail
      Contact( "R-201_Control_DB".FromHMI.Initialize )
      I_Contact( "R-201_Control_DB".FromHMI.Start )
      wire#w1
      I_Contact( "Control_Read_FROM_R-201_DB".Initialization_Done )
      Coil( "R-201_Control_DB".Cmds.Initialize )
   END_RUNG
   RUNG wire#powerrail
      Contact( "R-201_Control_DB".Cmds.Initialize )
   END_RUNG wire#w1
   // the same network as SCL:
   "R-201_Control_DB".Cmds.Initialize := (("R-201_Control_DB".FromHMI.Initialize AND NOT "R-201_Control_DB".FromHMI.Start) OR "R-201_Control_DB".Cmds.Initialize) AND NOT "Control_Read_FROM_R-201_DB".Initialization_Done;
END_REGION

REGION Network 5: Start
   RUNG wire#powerrail
      Contact( "R-201_Control_DB".FromHMI.Start )
      I_Contact( "R-201_Control_DB".FromHMI.Initialize )
      Coil( "R-201_Control_DB".Cmds.Start )
   END_RUNG
   // the same network as SCL:
   "R-201_Control_DB".Cmds.Start := "R-201_Control_DB".FromHMI.Start AND NOT "R-201_Control_DB".FromHMI.Initialize;
END_REGION

REGION Network 6: Tank Wash
   RUNG wire#powerrail
      Contact( "R-201_Control_DB".FromHMI.TankWash )
      I_Contact( "R-201_Control_DB".FromHMI.Start )
      Coil( "R-201_Control_DB".Cmds.TankWash )
   END_RUNG
   // the same network as SCL:
   "R-201_Control_DB".Cmds.TankWash := "R-201_Control_DB".FromHMI.TankWash AND NOT "R-201_Control_DB".FromHMI.Start;
END_REGION

REGION Network 7: Tube Wash
   RUNG wire#powerrail
      Contact( "R-201_Control_DB".FromHMI.TubeWash )
      I_Contact( "R-201_Control_DB".FromHMI.Start )
      Coil( "R-201_Control_DB".Cmds.TubeWash )
   END_RUNG
   // the same network as SCL:
   "R-201_Control_DB".Cmds.TubeWash := "R-201_Control_DB".FromHMI.TubeWash AND NOT "R-201_Control_DB".FromHMI.Start;
END_REGION
END_FUNCTION

// folder: State MACHINE/2)Reactors/Reactor R-201/Control R-201/Control <---> R-201

FUNCTION "Control_Signals_FROM_R-201" : Void   // FC45, LAD
{ S7_Optimized_Access := 'TRUE' }
VERSION : 0.1
BEGIN

REGION Network 1: R-201 Initialization Done
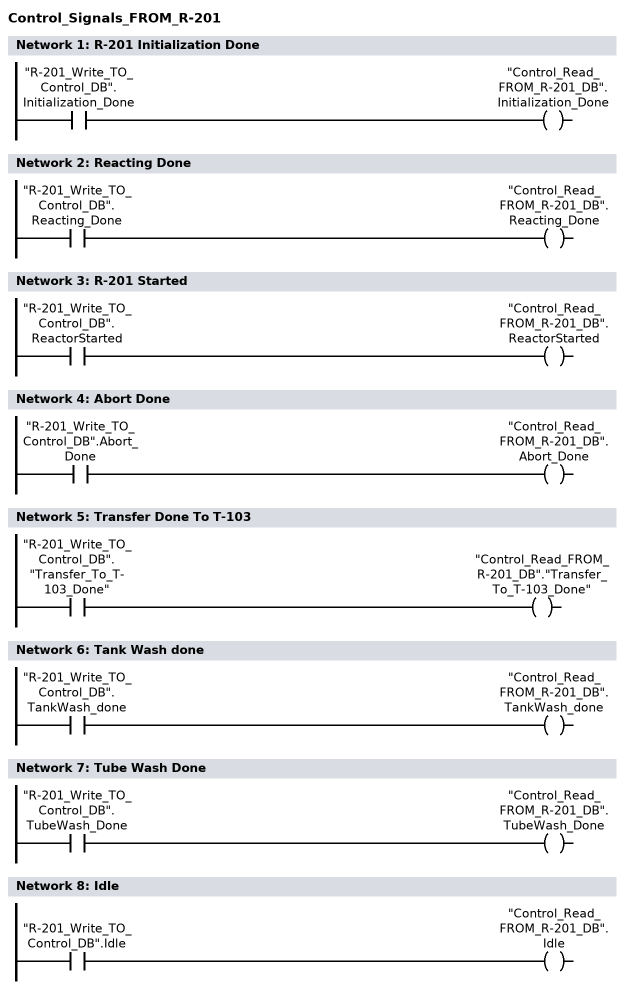
   RUNG wire#powerrail
      Contact( "R-201_Write_TO_Control_DB".Initialization_Done )
      Coil( "Control_Read_FROM_R-201_DB".Initialization_Done )
   END_RUNG
   // the same network as SCL:
   "Control_Read_FROM_R-201_DB".Initialization_Done := "R-201_Write_TO_Control_DB".Initialization_Done;
END_REGION

REGION Network 2: Reacting Done
   RUNG wire#powerrail
      Contact( "R-201_Write_TO_Control_DB".Reacting_Done )
      Coil( "Control_Read_FROM_R-201_DB".Reacting_Done )
   END_RUNG
   // the same network as SCL:
   "Control_Read_FROM_R-201_DB".Reacting_Done := "R-201_Write_TO_Control_DB".Reacting_Done;
END_REGION

REGION Network 3: R-201 Started
   RUNG wire#powerrail
      Contact( "R-201_Write_TO_Control_DB".ReactorStarted )
      Coil( "Control_Read_FROM_R-201_DB".ReactorStarted )
   END_RUNG
   // the same network as SCL:
   "Control_Read_FROM_R-201_DB".ReactorStarted := "R-201_Write_TO_Control_DB".ReactorStarted;
END_REGION

REGION Network 4: Abort Done
   RUNG wire#powerrail
      Contact( "R-201_Write_TO_Control_DB".Abort_Done )
      Coil( "Control_Read_FROM_R-201_DB".Abort_Done )
   END_RUNG
   // the same network as SCL:
   "Control_Read_FROM_R-201_DB".Abort_Done := "R-201_Write_TO_Control_DB".Abort_Done;
END_REGION
